REGION Network 333
   RUNG wire#powerrail
      Move(in := "DuplicateCarrierNumber", out1 => "Carrier_66_Duplicate_Carrier_Number")
   END_RUNG
   // the same network as SCL:
   "Carrier_66_Duplicate_Carrier_Number" := "DuplicateCarrierNumber";
END_REGION

REGION Network 334
   RUNG wire#powerrail
      Move(in := "FirstDuplicateCarrierPosition", out1 => "Carrier_66_First_Duplicate_Carrier_Position")
   END_RUNG
   // the same network as SCL:
   "Carrier_66_First_Duplicate_Carrier_Position" := "FirstDuplicateCarrierPosition";
END_REGION

REGION Network 335
   RUNG wire#powerrail
      Move(in := "SecondDuplicateCarrierPosition", out1 => "Carrier_66_Second_Duplicate_Carrier_Position")
   END_RUNG
   // the same network as SCL:
   "Carrier_66_Second_Duplicate_Carrier_Position" := "SecondDuplicateCarrierPosition";
END_REGION

REGION Network 336
   RUNG wire#powerrail
      Contact( "EMS".Carrier[66].SDC_OUT.HeartBeat )
      Coil( "Carrier_66_Heartbeat" )
   END_RUNG
   // the same network as SCL:
   "Carrier_66_Heartbeat" := "EMS".Carrier[66].SDC_OUT.HeartBeat;
END_REGION

REGION Network 337
   RUNG wire#powerrail
      Contact( "EMS".Carrier[66].SDC_OUT.DriveFwdCMD )
      I_Contact( "EMS".Carrier[65].SDC_IN.CrashDetectStatus )
      Coil( "Carrier_66_Drive_Forward_Command" )
   END_RUNG
   // the same network as SCL:
   "Carrier_66_Drive_Forward_Command" := "EMS".Carrier[66].SDC_OUT.DriveFwdCMD AND NOT "EMS".Carrier[65].SDC_IN.CrashDetectStatus;
END_REGION

REGION Network 338
   RUNG wire#powerrail
      Contact( "EMS".Carrier[66].SDC_OUT.FaultReset )
      Coil( "Carrier_66_Fault_Reset" )
   END_RUNG
   // the same network as SCL:
   "Carrier_66_Fault_Reset" := "EMS".Carrier[66].SDC_OUT.FaultReset;
END_REGION

REGION Network 339
   RUNG wire#powerrail
      Contact( "EMS".Carrier[66].SDC_OUT.AtCmdPos )
      Coil( "Carrier_66_At_Command_Position" )
   END_RUNG
   // the same network as SCL:
   "Carrier_66_At_Command_Position" := "EMS".Carrier[66].SDC_OUT.AtCmdPos;
END_REGION

REGION Network 340
   RUNG wire#powerrail
      Contact( "DuplicateCarrierfound" )
      Coil( "Carrier_66_Duplicate_Carrier_Fault" )
   END_RUNG
   // the same network as SCL:
   "Carrier_66_Duplicate_Carrier_Fault" := "DuplicateCarrierfound";
END_REGION

REGION Network 341
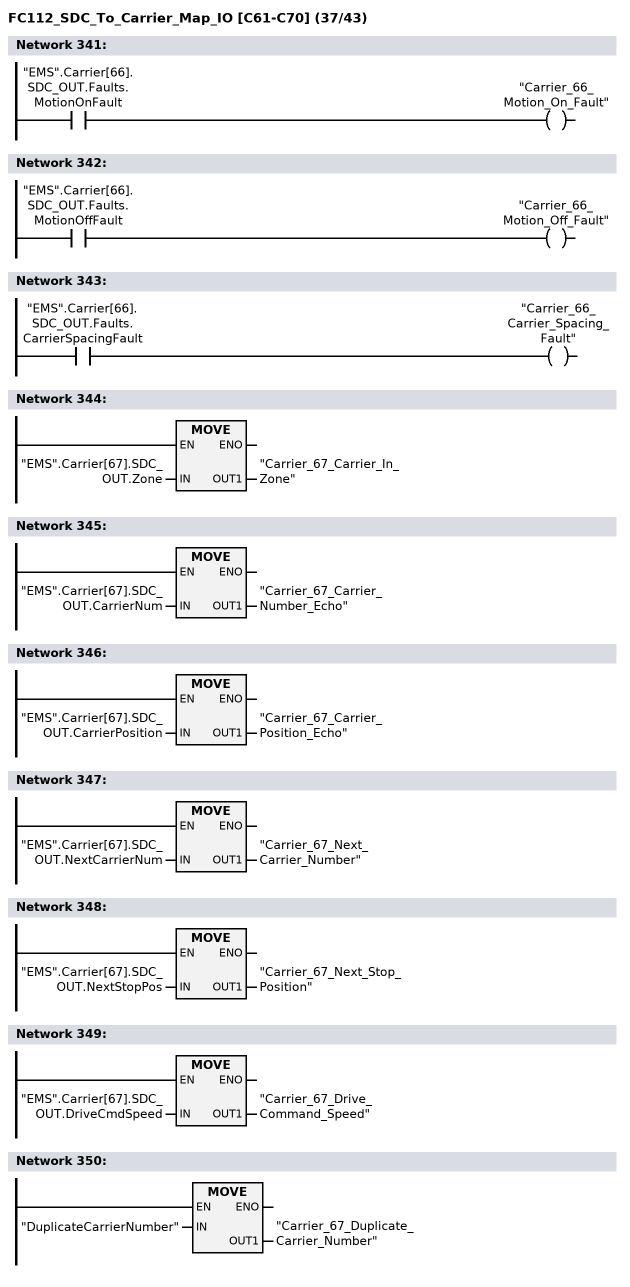
   RUNG wire#powerrail
      Contact( "EMS".Carrier[66].SDC_OUT.Faults.MotionOnFault )
      Coil( "Carrier_66_Motion_On_Fault" )
   END_RUNG
   // the same network as SCL:
   "Carrier_66_Motion_On_Fault" := "EMS".Carrier[66].SDC_OUT.Faults.MotionOnFault;
END_REGION

REGION Network 342
   RUNG wire#powerrail
      Contact( "EMS".Carrier[66].SDC_OUT.Faults.MotionOffFault )
      Coil( "Carrier_66_Motion_Off_Fault" )
   END_RUNG
   // the same network as SCL:
   "Carrier_66_Motion_Off_Fault" := "EMS".Carrier[66].SDC_OUT.Faults.MotionOffFault;
END_REGION

REGION Network 343
   RUNG wire#powerrail
      Contact( "EMS".Carrier[66].SDC_OUT.Faults.CarrierSpacingFault )
      Coil( "Carrier_66_Carrier_Spacing_Fault" )
   END_RUNG
   // the same network as SCL:
   "Carrier_66_Carrier_Spacing_Fault" := "EMS".Carrier[66].SDC_OUT.Faults.CarrierSpacingFault;
END_REGION

REGION Network 344
   RUNG wire#powerrail
      Move(in := "EMS".Carrier[67].SDC_OUT.Zone, out1 => "Carrier_67_Carrier_In_Zone")
   END_RUNG
   // the same network as SCL:
   "Carrier_67_Carrier_In_Zone" := "EMS".Carrier[67].SDC_OUT.Zone;
END_REGION

REGION Network 345
   RUNG wire#powerrail
      Move(in := "EMS".Carrier[67].SDC_OUT.CarrierNum, out1 => "Carrier_67_Carrier_Number_Echo")
   END_RUNG
   // the same network as SCL:
   "Carrier_67_Carrier_Number_Echo" := "EMS".Carrier[67].SDC_OUT.CarrierNum;
END_REGION

REGION Network 346
   RUNG wire#powerrail
      Move(in := "EMS".Carrier[67].SDC_OUT.CarrierPosition, out1 => "Carrier_67_Carrier_Position_Echo")
   END_RUNG
   // the same network as SCL:
   "Carrier_67_Carrier_Position_Echo" := "EMS".Carrier[67].SDC_OUT.CarrierPosition;
END_REGION

REGION Network 347
   RUNG wire#powerrail
      Move(in := "EMS".Carrier[67].SDC_OUT.NextCarrierNum, out1 => "Carrier_67_Next_Carrier_Number")
   END_RUNG
   // the same network as SCL:
   "Carrier_67_Next_Carrier_Number" := "EMS".Carrier[67].SDC_OUT.NextCarrierNum;
END_REGION

REGION Network 348
   RUNG wire#powerrail
      Move(in := "EMS".Carrier[67].SDC_OUT.NextStopPos, out1 => "Carrier_67_Next_Stop_Position")
   END_RUNG
   // the same network as SCL:
   "Carrier_67_Next_Stop_Position" := "EMS".Carrier[67].SDC_OUT.NextStopPos;
END_REGION

REGION Network 349
   RUNG wire#powerrail
      Move(in := "EMS".Carrier[67].SDC_OUT.DriveCmdSpeed, out1 => "Carrier_67_Drive_Command_Speed")
   END_RUNG
   // the same network as SCL:
   "Carrier_67_Drive_Command_Speed" := "EMS".Carrier[67].SDC_OUT.DriveCmdSpeed;
END_REGION

REGION Network 350
   RUNG wire#powerrail
      Move(in := "DuplicateCarrierNumber", out1 => "Carrier_67_Duplicate_Carrier_Number")
   END_RUNG
   // the same network as SCL:
   "Carrier_67_Duplicate_Carrier_Number" := "DuplicateCarrierNumber";
END_REGION

REGION Network 351
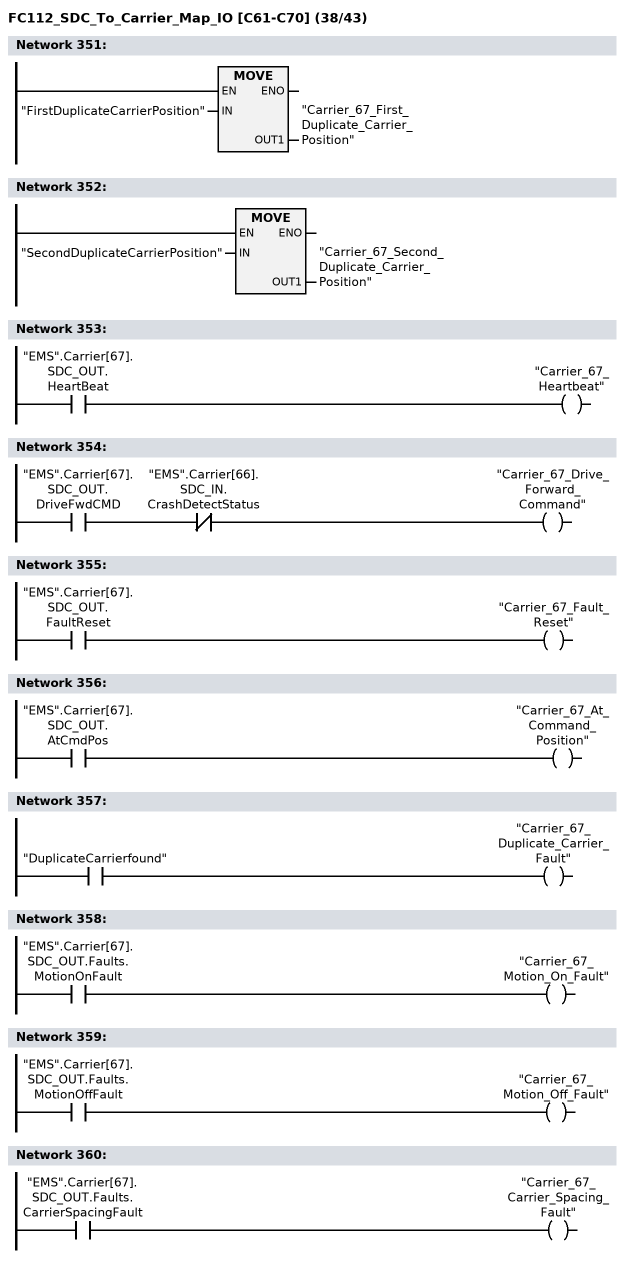
   RUNG wire#powerrail
      Move(in := "FirstDuplicateCarrierPosition", out1 => "Carrier_67_First_Duplicate_Carrier_Position")
   END_RUNG
   // the same network as SCL:
   "Carrier_67_First_Duplicate_Carrier_Position" := "FirstDuplicateCarrierPosition";
END_REGION

REGION Network 352
   RUNG wire#powerrail
      Move(in := "SecondDuplicateCarrierPosition", out1 => "Carrier_67_Second_Duplicate_Carrier_Position")
   END_RUNG
   // the same network as SCL:
   "Carrier_67_Second_Duplicate_Carrier_Position" := "SecondDuplicateCarrierPosition";
END_REGION

REGION Network 353
   RUNG wire#powerrail
      Contact( "EMS".Carrier[67].SDC_OUT.HeartBeat )
      Coil( "Carrier_67_Heartbeat" )
   END_RUNG
   // the same network as SCL:
   "Carrier_67_Heartbeat" := "EMS".Carrier[67].SDC_OUT.HeartBeat;
END_REGION

REGION Network 354
   RUNG wire#powerrail
      Contact( "EMS".Carrier[67].SDC_OUT.DriveFwdCMD )
      I_Contact( "EMS".Carrier[66].SDC_IN.CrashDetectStatus )
      Coil( "Carrier_67_Drive_Forward_Command" )
   END_RUNG
   // the same network as SCL:
   "Carrier_67_Drive_Forward_Command" := "EMS".Carrier[67].SDC_OUT.DriveFwdCMD AND NOT "EMS".Carrier[66].SDC_IN.CrashDetectStatus;
END_REGION

REGION Network 355
   RUNG wire#powerrail
      Contact( "EMS".Carrier[67].SDC_OUT.FaultReset )
      Coil( "Carrier_67_Fault_Reset" )
   END_RUNG
   // the same network as SCL:
   "Carrier_67_Fault_Reset" := "EMS".Carrier[67].SDC_OUT.FaultReset;
END_REGION

REGION Network 356
   RUNG wire#powerrail
      Contact( "EMS".Carrier[67].SDC_OUT.AtCmdPos )
      Coil( "Carrier_67_At_Command_Position" )
   END_RUNG
   // the same network as SCL:
   "Carrier_67_At_Command_Position" := "EMS".Carrier[67].SDC_OUT.AtCmdPos;
END_REGION

REGION Network 357
   RUNG wire#powerrail
      Contact( "DuplicateCarrierfound" )
      Coil( "Carrier_67_Duplicate_Carrier_Fault" )
   END_RUNG
   // the same network as SCL:
   "Carrier_67_Duplicate_Carrier_Fault" := "DuplicateCarrierfound";
END_REGION

REGION Network 358
   RUNG wire#powerrail
      Contact( "EMS".Carrier[67].SDC_OUT.Faults.MotionOnFault )
      Coil( "Carrier_67_Motion_On_Fault" )
   END_RUNG
   // the same network as SCL:
   "Carrier_67_Motion_On_Fault" := "EMS".Carrier[67].SDC_OUT.Faults.MotionOnFault;
END_REGION

REGION Network 359
   RUNG wire#powerrail
      Contact( "EMS".Carrier[67].SDC_OUT.Faults.MotionOffFault )
      Coil( "Carrier_67_Motion_Off_Fault" )
   END_RUNG
   // the same network as SCL:
   "Carrier_67_Motion_Off_Fault" := "EMS".Carrier[67].SDC_OUT.Faults.MotionOffFault;
END_REGION

REGION Network 360
   RUNG wire#powerrail
      Contact( "EMS".Carrier[67].SDC_OUT.Faults.CarrierSpacingFault )
      Coil( "Carrier_67_Carrier_Spacing_Fault" )
   END_RUNG
   // the same network as SCL:
   "Carrier_67_Carrier_Spacing_Fault" := "EMS".Carrier[67].SDC_OUT.Faults.CarrierSpacingFault;
END_REGION

REGION Network 361
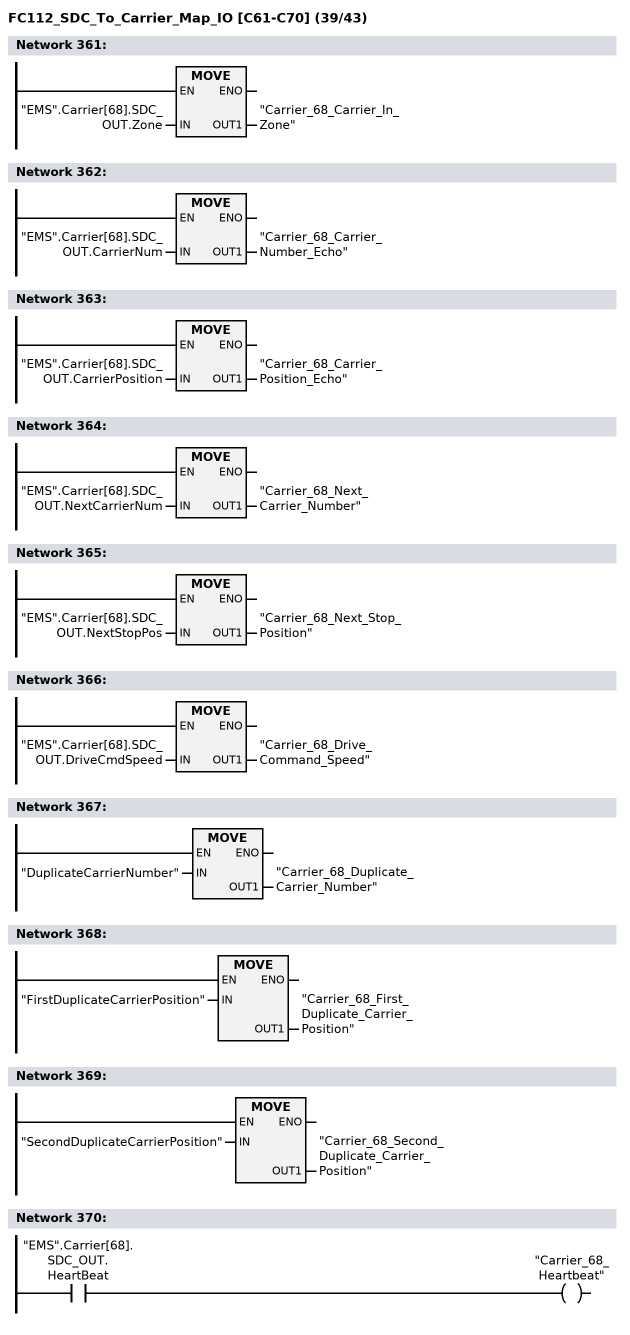
   RUNG wire#powerrail
      Move(in := "EMS".Carrier[68].SDC_OUT.Zone, out1 => "Carrier_68_Carrier_In_Zone")
   END_RUNG
   // the same network as SCL:
   "Carrier_68_Carrier_In_Zone" := "EMS".Carrier[68].SDC_OUT.Zone;
END_REGION

REGION Network 362
   RUNG wire#powerrail
      Move(in := "EMS".Carrier[68].SDC_OUT.CarrierNum, out1 => "Carrier_68_Carrier_Number_Echo")
   END_RUNG
   // the same network as SCL:
   "Carrier_68_Carrier_Number_Echo" := "EMS".Carrier[68].SDC_OUT.CarrierNum;
END_REGION

REGION Network 363
   RUNG wire#powerrail
      Move(in := "EMS".Carrier[68].SDC_OUT.CarrierPosition, out1 => "Carrier_68_Carrier_Position_Echo")
   END_RUNG
   // the same network as SCL:
   "Carrier_68_Carrier_Position_Echo" := "EMS".Carrier[68].SDC_OUT.CarrierPosition;
END_REGION

REGION Network 364
   RUNG wire#powerrail
      Move(in := "EMS".Carrier[68].SDC_OUT.NextCarrierNum, out1 => "Carrier_68_Next_Carrier_Number")
   END_RUNG
   // the same network as SCL:
   "Carrier_68_Next_Carrier_Number" := "EMS".Carrier[68].SDC_OUT.NextCarrierNum;
END_REGION

REGION Network 365
   RUNG wire#powerrail
      Move(in := "EMS".Carrier[68].SDC_OUT.NextStopPos, out1 => "Carrier_68_Next_Stop_Position")
   END_RUNG
   // the same network as SCL:
   "Carrier_68_Next_Stop_Position" := "EMS".Carrier[68].SDC_OUT.NextStopPos;
END_REGION

REGION Network 366
   RUNG wire#powerrail
      Move(in := "EMS".Carrier[68].SDC_OUT.DriveCmdSpeed, out1 => "Carrier_68_Drive_Command_Speed")
   END_RUNG
   // the same network as SCL:
   "Carrier_68_Drive_Command_Speed" := "EMS".Carrier[68].SDC_OUT.DriveCmdSpeed;
END_REGION

REGION Network 367
   RUNG wire#powerrail
      Move(in := "DuplicateCarrierNumber", out1 => "Carrier_68_Duplicate_Carrier_Number")
   END_RUNG
   // the same network as SCL:
   "Carrier_68_Duplicate_Carrier_Number" := "DuplicateCarrierNumber";
END_REGION

REGION Network 368
   RUNG wire#powerrail
      Move(in := "FirstDuplicateCarrierPosition", out1 => "Carrier_68_First_Duplicate_Carrier_Position")
   END_RUNG
   // the same network as SCL:
   "Carrier_68_First_Duplicate_Carrier_Position" := "FirstDuplicateCarrierPosition";
END_REGION

REGION Network 369
   RUNG wire#powerrail
      Move(in := "SecondDuplicateCarrierPosition", out1 => "Carrier_68_Second_Duplicate_Carrier_Position")
   END_RUNG
   // the same network as SCL:
   "Carrier_68_Second_Duplicate_Carrier_Position" := "SecondDuplicateCarrierPosition";
END_REGION

REGION Network 370
   RUNG wire#powerrail
      Contact( "EMS".Carrier[68].SDC_OUT.HeartBeat )
      Coil( "Carrier_68_Heartbeat" )
   END_RUNG
   // the same network as SCL:
   "Carrier_68_Heartbeat" := "EMS".Carrier[68].SDC_OUT.HeartBeat;
END_REGION

REGION Network 371
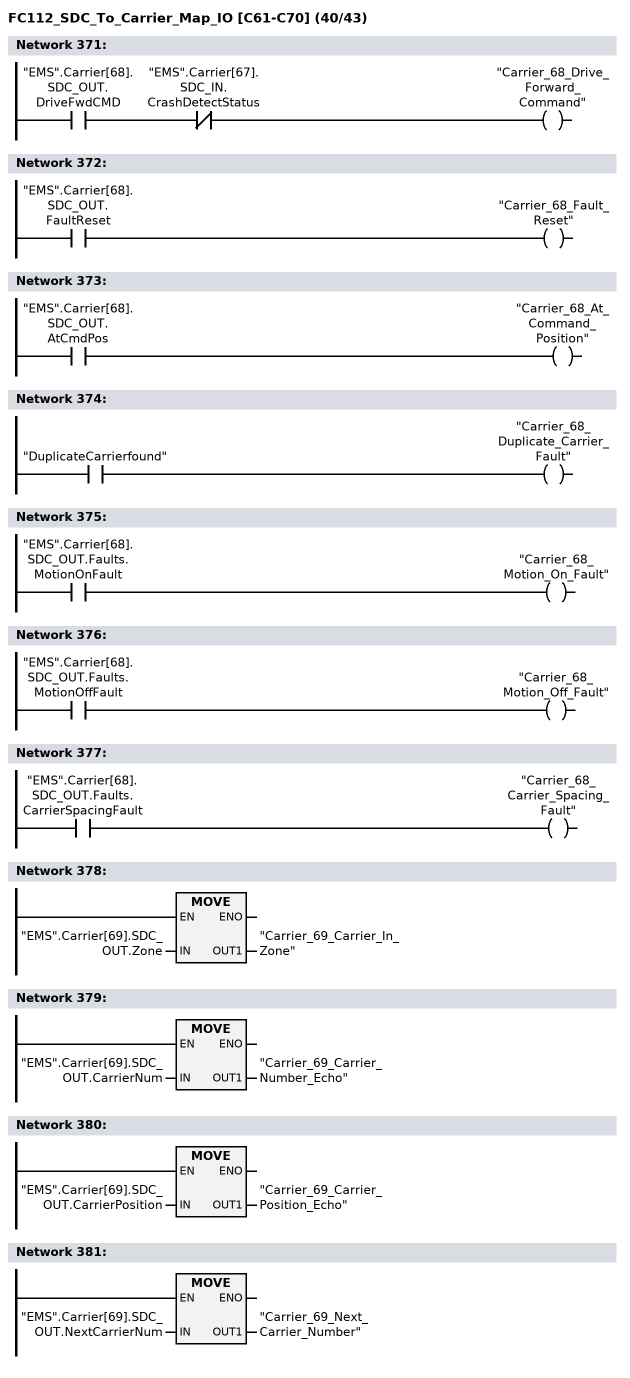
   RUNG wire#powerrail
      Contact( "EMS".Carrier[68].SDC_OUT.DriveFwdCMD )
      I_Contact( "EMS".Carrier[67].SDC_IN.CrashDetectStatus )
      Coil( "Carrier_68_Drive_Forward_Command" )
   END_RUNG
   // the same network as SCL:
   "Carrier_68_Drive_Forward_Command" := "EMS".Carrier[68].SDC_OUT.DriveFwdCMD AND NOT "EMS".Carrier[67].SDC_IN.CrashDetectStatus;
END_REGION

REGION Network 372
   RUNG wire#powerrail
      Contact( "EMS".Carrier[68].SDC_OUT.FaultReset )
      Coil( "Carrier_68_Fault_Reset" )
   END_RUNG
   // the same network as SCL:
   "Carrier_68_Fault_Reset" := "EMS".Carrier[68].SDC_OUT.FaultReset;
END_REGION

REGION Network 373
   RUNG wire#powerrail
      Contact( "EMS".Carrier[68].SDC_OUT.AtCmdPos )
      Coil( "Carrier_68_At_Command_Position" )
   END_RUNG
   // the same network as SCL:
   "Carrier_68_At_Command_Position" := "EMS".Carrier[68].SDC_OUT.AtCmdPos;
END_REGION

REGION Network 374
   RUNG wire#powerrail
      Contact( "DuplicateCarrierfound" )
      Coil( "Carrier_68_Duplicate_Carrier_Fault" )
   END_RUNG
   // the same network as SCL:
   "Carrier_68_Duplicate_Carrier_Fault" := "DuplicateCarrierfound";
END_REGION

REGION Network 375
   RUNG wire#powerrail
      Contact( "EMS".Carrier[68].SDC_OUT.Faults.MotionOnFault )
      Coil( "Carrier_68_Motion_On_Fault" )
   END_RUNG
   // the same network as SCL:
   "Carrier_68_Motion_On_Fault" := "EMS".Carrier[68].SDC_OUT.Faults.MotionOnFault;
END_REGION

REGION Network 376
   RUNG wire#powerrail
      Contact( "EMS".Carrier[68].SDC_OUT.Faults.MotionOffFault )
      Coil( "Carrier_68_Motion_Off_Fault" )
   END_RUNG
   // the same network as SCL:
   "Carrier_68_Motion_Off_Fault" := "EMS".Carrier[68].SDC_OUT.Faults.MotionOffFault;
END_REGION

REGION Network 377
   RUNG wire#powerrail
      Contact( "EMS".Carrier[68].SDC_OUT.Faults.CarrierSpacingFault )
      Coil( "Carrier_68_Carrier_Spacing_Fault" )
   END_RUNG
   // the same network as SCL:
   "Carrier_68_Carrier_Spacing_Fault" := "EMS".Carrier[68].SDC_OUT.Faults.CarrierSpacingFault;
END_REGION

REGION Network 378
   RUNG wire#powerrail
      Move(in := "EMS".Carrier[69].SDC_OUT.Zone, out1 => "Carrier_69_Carrier_In_Zone")
   END_RUNG
   // the same network as SCL:
   "Carrier_69_Carrier_In_Zone" := "EMS".Carrier[69].SDC_OUT.Zone;
END_REGION

REGION Network 379
   RUNG wire#powerrail
      Move(in := "EMS".Carrier[69].SDC_OUT.CarrierNum, out1 => "Carrier_69_Carrier_Number_Echo")
   END_RUNG
   // the same network as SCL:
   "Carrier_69_Carrier_Number_Echo" := "EMS".Carrier[69].SDC_OUT.CarrierNum;
END_REGION

REGION Network 380
   RUNG wire#powerrail
      Move(in := "EMS".Carrier[69].SDC_OUT.CarrierPosition, out1 => "Carrier_69_Carrier_Position_Echo")
   END_RUNG
   // the same network as SCL:
   "Carrier_69_Carrier_Position_Echo" := "EMS".Carrier[69].SDC_OUT.CarrierPosition;
END_REGION

REGION Network 381
   RUNG wire#powerrail
      Move(in := "EMS".Carrier[69].SDC_OUT.NextCarrierNum, out1 => "Carrier_69_Next_Carrier_Number")
   END_RUNG
   // the same network as SCL:
   "Carrier_69_Next_Carrier_Number" := "EMS".Carrier[69].SDC_OUT.NextCarrierNum;
END_REGION

REGION Network 382
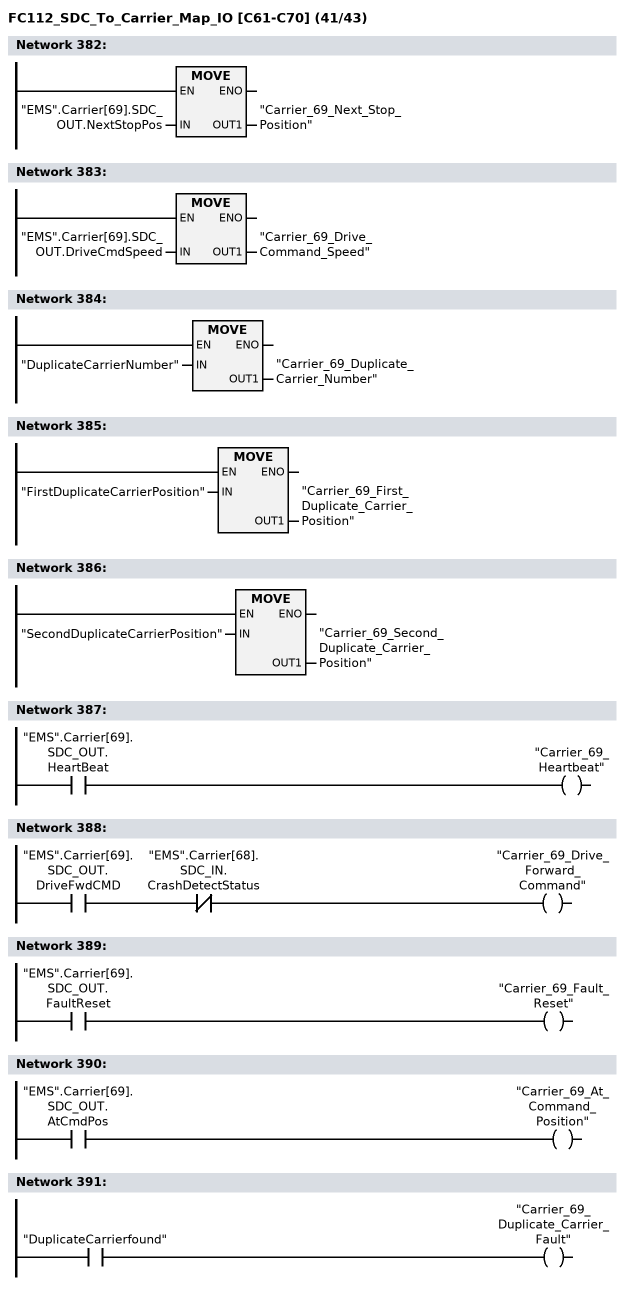
   RUNG wire#powerrail
      Move(in := "EMS".Carrier[69].SDC_OUT.NextStopPos, out1 => "Carrier_69_Next_Stop_Position")
   END_RUNG
   // the same network as SCL:
   "Carrier_69_Next_Stop_Position" := "EMS".Carrier[69].SDC_OUT.NextStopPos;
END_REGION

REGION Network 383
   RUNG wire#powerrail
      Move(in := "EMS".Carrier[69].SDC_OUT.DriveCmdSpeed, out1 => "Carrier_69_Drive_Command_Speed")
   END_RUNG
   // the same network as SCL:
   "Carrier_69_Drive_Command_Speed" := "EMS".Carrier[69].SDC_OUT.DriveCmdSpeed;
END_REGION

REGION Network 384
   RUNG wire#powerrail
      Move(in := "DuplicateCarrierNumber", out1 => "Carrier_69_Duplicate_Carrier_Number")
   END_RUNG
   // the same network as SCL:
   "Carrier_69_Duplicate_Carrier_Number" := "DuplicateCarrierNumber";
END_REGION

REGION Network 385
   RUNG wire#powerrail
      Move(in := "FirstDuplicateCarrierPosition", out1 => "Carrier_69_First_Duplicate_Carrier_Position")
   END_RUNG
   // the same network as SCL:
   "Carrier_69_First_Duplicate_Carrier_Position" := "FirstDuplicateCarrierPosition";
END_REGION

REGION Network 386
   RUNG wire#powerrail
      Move(in := "SecondDuplicateCarrierPosition", out1 => "Carrier_69_Second_Duplicate_Carrier_Position")
   END_RUNG
   // the same network as SCL:
   "Carrier_69_Second_Duplicate_Carrier_Position" := "SecondDuplicateCarrierPosition";
END_REGION

REGION Network 387
   RUNG wire#powerrail
      Contact( "EMS".Carrier[69].SDC_OUT.HeartBeat )
      Coil( "Carrier_69_Heartbeat" )
   END_RUNG
   // the same network as SCL:
   "Carrier_69_Heartbeat" := "EMS".Carrier[69].SDC_OUT.HeartBeat;
END_REGION

REGION Network 388
   RUNG wire#powerrail
      Contact( "EMS".Carrier[69].SDC_OUT.DriveFwdCMD )
      I_Contact( "EMS".Carrier[68].SDC_IN.CrashDetectStatus )
      Coil( "Carrier_69_Drive_Forward_Command" )
   END_RUNG
   // the same network as SCL:
   "Carrier_69_Drive_Forward_Command" := "EMS".Carrier[69].SDC_OUT.DriveFwdCMD AND NOT "EMS".Carrier[68].SDC_IN.CrashDetectStatus;
END_REGION

REGION Network 389
   RUNG wire#powerrail
      Contact( "EMS".Carrier[69].SDC_OUT.FaultReset )
      Coil( "Carrier_69_Fault_Reset" )
   END_RUNG
   // the same network as SCL:
   "Carrier_69_Fault_Reset" := "EMS".Carrier[69].SDC_OUT.FaultReset;
END_REGION

REGION Network 390
   RUNG wire#powerrail
      Contact( "EMS".Carrier[69].SDC_OUT.AtCmdPos )
      Coil( "Carrier_69_At_Command_Position" )
   END_RUNG
   // the same network as SCL:
   "Carrier_69_At_Command_Position" := "EMS".Carrier[69].SDC_OUT.AtCmdPos;
END_REGION

REGION Network 391
   RUNG wire#powerrail
      Contact( "DuplicateCarrierfound" )
      Coil( "Carrier_69_Duplicate_Carrier_Fault" )
   END_RUNG
   // the same network as SCL:
   "Carrier_69_Duplicate_Carrier_Fault" := "DuplicateCarrierfound";
END_REGION

REGION Network 392
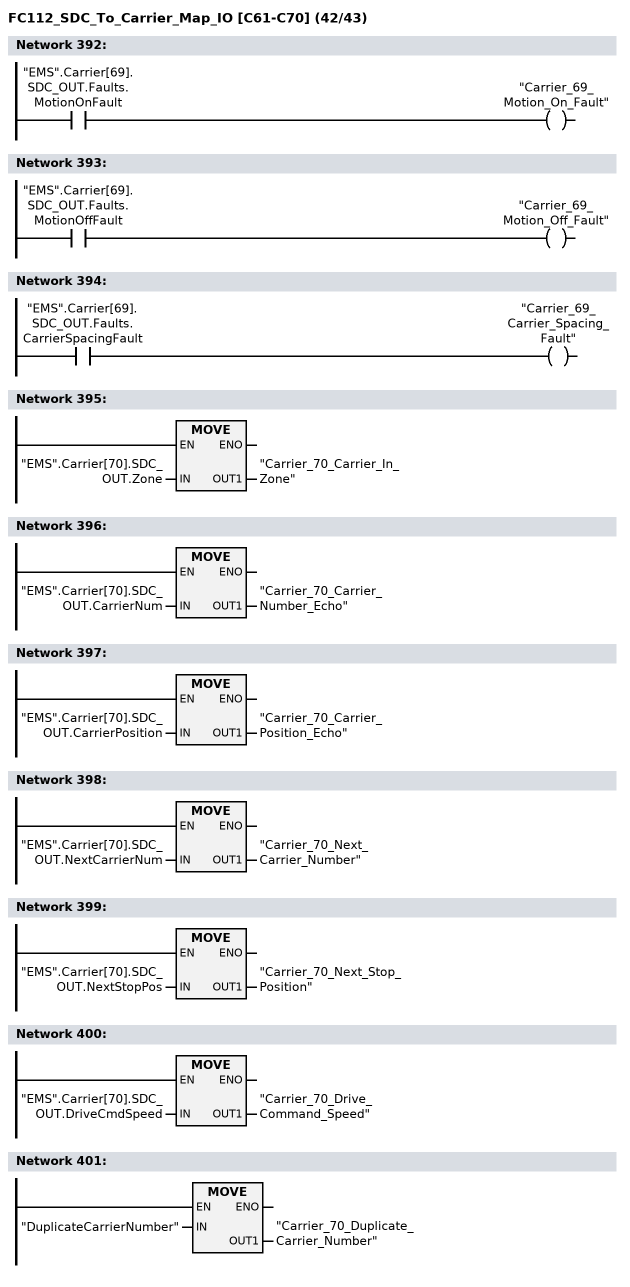
   RUNG wire#powerrail
      Contact( "EMS".Carrier[69].SDC_OUT.Faults.MotionOnFault )
      Coil( "Carrier_69_Motion_On_Fault" )
   END_RUNG
   // the same network as SCL:
   "Carrier_69_Motion_On_Fault" := "EMS".Carrier[69].SDC_OUT.Faults.MotionOnFault;
END_REGION

REGION Network 393
   RUNG wire#powerrail
      Contact( "EMS".Carrier[69].SDC_OUT.Faults.MotionOffFault )
      Coil( "Carrier_69_Motion_Off_Fault" )
   END_RUNG
   // the same network as SCL:
   "Carrier_69_Motion_Off_Fault" := "EMS".Carrier[69].SDC_OUT.Faults.MotionOffFault;
END_REGION

REGION Network 394
   RUNG wire#powerrail
      Contact( "EMS".Carrier[69].SDC_OUT.Faults.CarrierSpacingFault )
      Coil( "Carrier_69_Carrier_Spacing_Fault" )
   END_RUNG
   // the same network as SCL:
   "Carrier_69_Carrier_Spacing_Fault" := "EMS".Carrier[69].SDC_OUT.Faults.CarrierSpacingFault;
END_REGION

REGION Network 395
   RUNG wire#powerrail
      Move(in := "EMS".Carrier[70].SDC_OUT.Zone, out1 => "Carrier_70_Carrier_In_Zone")
   END_RUNG
   // the same network as SCL:
   "Carrier_70_Carrier_In_Zone" := "EMS".Carrier[70].SDC_OUT.Zone;
END_REGION

REGION Network 396
   RUNG wire#powerrail
      Move(in := "EMS".Carrier[70].SDC_OUT.CarrierNum, out1 => "Carrier_70_Carrier_Number_Echo")
   END_RUNG
   // the same network as SCL:
   "Carrier_70_Carrier_Number_Echo" := "EMS".Carrier[70].SDC_OUT.CarrierNum;
END_REGION

REGION Network 397
   RUNG wire#powerrail
      Move(in := "EMS".Carrier[70].SDC_OUT.CarrierPosition, out1 => "Carrier_70_Carrier_Position_Echo")
   END_RUNG
   // the same network as SCL:
   "Carrier_70_Carrier_Position_Echo" := "EMS".Carrier[70].SDC_OUT.CarrierPosition;
END_REGION

REGION Network 398
   RUNG wire#powerrail
      Move(in := "EMS".Carrier[70].SDC_OUT.NextCarrierNum, out1 => "Carrier_70_Next_Carrier_Number")
   END_RUNG
   // the same network as SCL:
   "Carrier_70_Next_Carrier_Number" := "EMS".Carrier[70].SDC_OUT.NextCarrierNum;
END_REGION

REGION Network 399
   RUNG wire#powerrail
      Move(in := "EMS".Carrier[70].SDC_OUT.NextStopPos, out1 => "Carrier_70_Next_Stop_Position")
   END_RUNG
   // the same network as SCL:
   "Carrier_70_Next_Stop_Position" := "EMS".Carrier[70].SDC_OUT.NextStopPos;
END_REGION

REGION Network 400
   RUNG wire#powerrail
      Move(in := "EMS".Carrier[70].SDC_OUT.DriveCmdSpeed, out1 => "Carrier_70_Drive_Command_Speed")
   END_RUNG
   // the same network as SCL:
   "Carrier_70_Drive_Command_Speed" := "EMS".Carrier[70].SDC_OUT.DriveCmdSpeed;
END_REGION

REGION Network 401
   RUNG wire#powerrail
      Move(in := "DuplicateCarrierNumber", out1 => "Carrier_70_Duplicate_Carrier_Number")
   END_RUNG
   // the same network as SCL:
   "Carrier_70_Duplicate_Carrier_Number" := "DuplicateCarrierNumber";
END_REGION

REGION Network 402
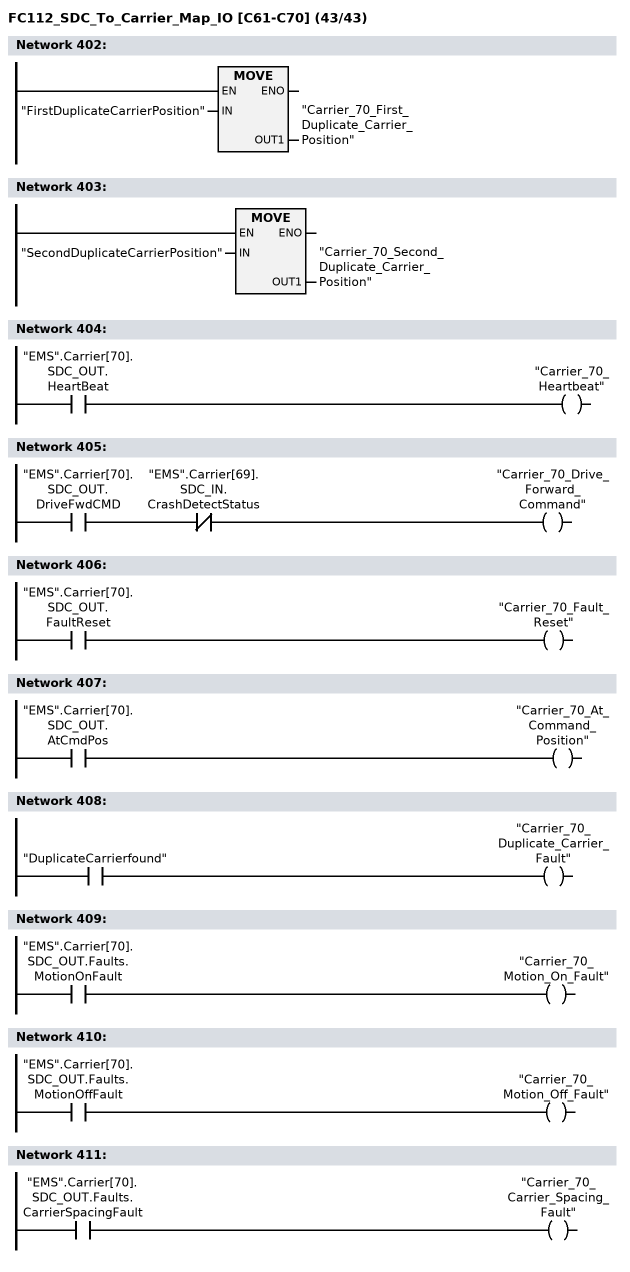
   RUNG wire#powerrail
      Move(in := "FirstDuplicateCarrierPosition", out1 => "Carrier_70_First_Duplicate_Carrier_Position")
   END_RUNG
   // the same network as SCL:
   "Carrier_70_First_Duplicate_Carrier_Position" := "FirstDuplicateCarrierPosition";
END_REGION

REGION Network 403
   RUNG wire#powerrail
      Move(in := "SecondDuplicateCarrierPosition", out1 => "Carrier_70_Second_Duplicate_Carrier_Position")
   END_RUNG
   // the same network as SCL:
   "Carrier_70_Second_Duplicate_Carrier_Position" := "SecondDuplicateCarrierPosition";
END_REGION

REGION Network 404
   RUNG wire#powerrail
      Contact( "EMS".Carrier[70].SDC_OUT.HeartBeat )
      Coil( "Carrier_70_Heartbeat" )
   END_RUNG
   // the same network as SCL:
   "Carrier_70_Heartbeat" := "EMS".Carrier[70].SDC_OUT.HeartBeat;
END_REGION

REGION Network 405
   RUNG wire#powerrail
      Contact( "EMS".Carrier[70].SDC_OUT.DriveFwdCMD )
      I_Contact( "EMS".Carrier[69].SDC_IN.CrashDetectStatus )
      Coil( "Carrier_70_Drive_Forward_Command" )
   END_RUNG
   // the same network as SCL:
   "Carrier_70_Drive_Forward_Command" := "EMS".Carrier[70].SDC_OUT.DriveFwdCMD AND NOT "EMS".Carrier[69].SDC_IN.CrashDetectStatus;
END_REGION

REGION Network 406
   RUNG wire#powerrail
      Contact( "EMS".Carrier[70].SDC_OUT.FaultReset )
      Coil( "Carrier_70_Fault_Reset" )
   END_RUNG
   // the same network as SCL:
   "Carrier_70_Fault_Reset" := "EMS".Carrier[70].SDC_OUT.FaultReset;
END_REGION

REGION Network 407
   RUNG wire#powerrail
      Contact( "EMS".Carrier[70].SDC_OUT.AtCmdPos )
      Coil( "Carrier_70_At_Command_Position" )
   END_RUNG
   // the same network as SCL:
   "Carrier_70_At_Command_Position" := "EMS".Carrier[70].SDC_OUT.AtCmdPos;
END_REGION

REGION Network 408
   RUNG wire#powerrail
      Contact( "DuplicateCarrierfound" )
      Coil( "Carrier_70_Duplicate_Carrier_Fault" )
   END_RUNG
   // the same network as SCL:
   "Carrier_70_Duplicate_Carrier_Fault" := "DuplicateCarrierfound";
END_REGION

REGION Network 409
   RUNG wire#powerrail
      Contact( "EMS".Carrier[70].SDC_OUT.Faults.MotionOnFault )
      Coil( "Carrier_70_Motion_On_Fault" )
   END_RUNG
   // the same network as SCL:
   "Carrier_70_Motion_On_Fault" := "EMS".Carrier[70].SDC_OUT.Faults.MotionOnFault;
END_REGION

REGION Network 410
   RUNG wire#powerrail
      Contact( "EMS".Carrier[70].SDC_OUT.Faults.MotionOffFault )
      Coil( "Carrier_70_Motion_Off_Fault" )
   END_RUNG
   // the same network as SCL:
   "Carrier_70_Motion_Off_Fault" := "EMS".Carrier[70].SDC_OUT.Faults.MotionOffFault;
END_REGION

REGION Network 411
   RUNG wire#powerrail
      Contact( "EMS".Carrier[70].SDC_OUT.Faults.CarrierSpacingFault )
      Coil( "Carrier_70_Carrier_Spacing_Fault" )
   END_RUNG
   // the same network as SCL:
   "Carrier_70_Carrier_Spacing_Fault" := "EMS".Carrier[70].SDC_OUT.Faults.CarrierSpacingFault;
END_REGION
END_FUNCTION

FUNCTION "FC113_SDC_To_Carrier_Map_IO [C71-C80]" : Void   // FC113, LAD
{ S7_Optimized_Access := 'TRUE' }
VERSION : 0.1
BEGIN

REGION Network 1
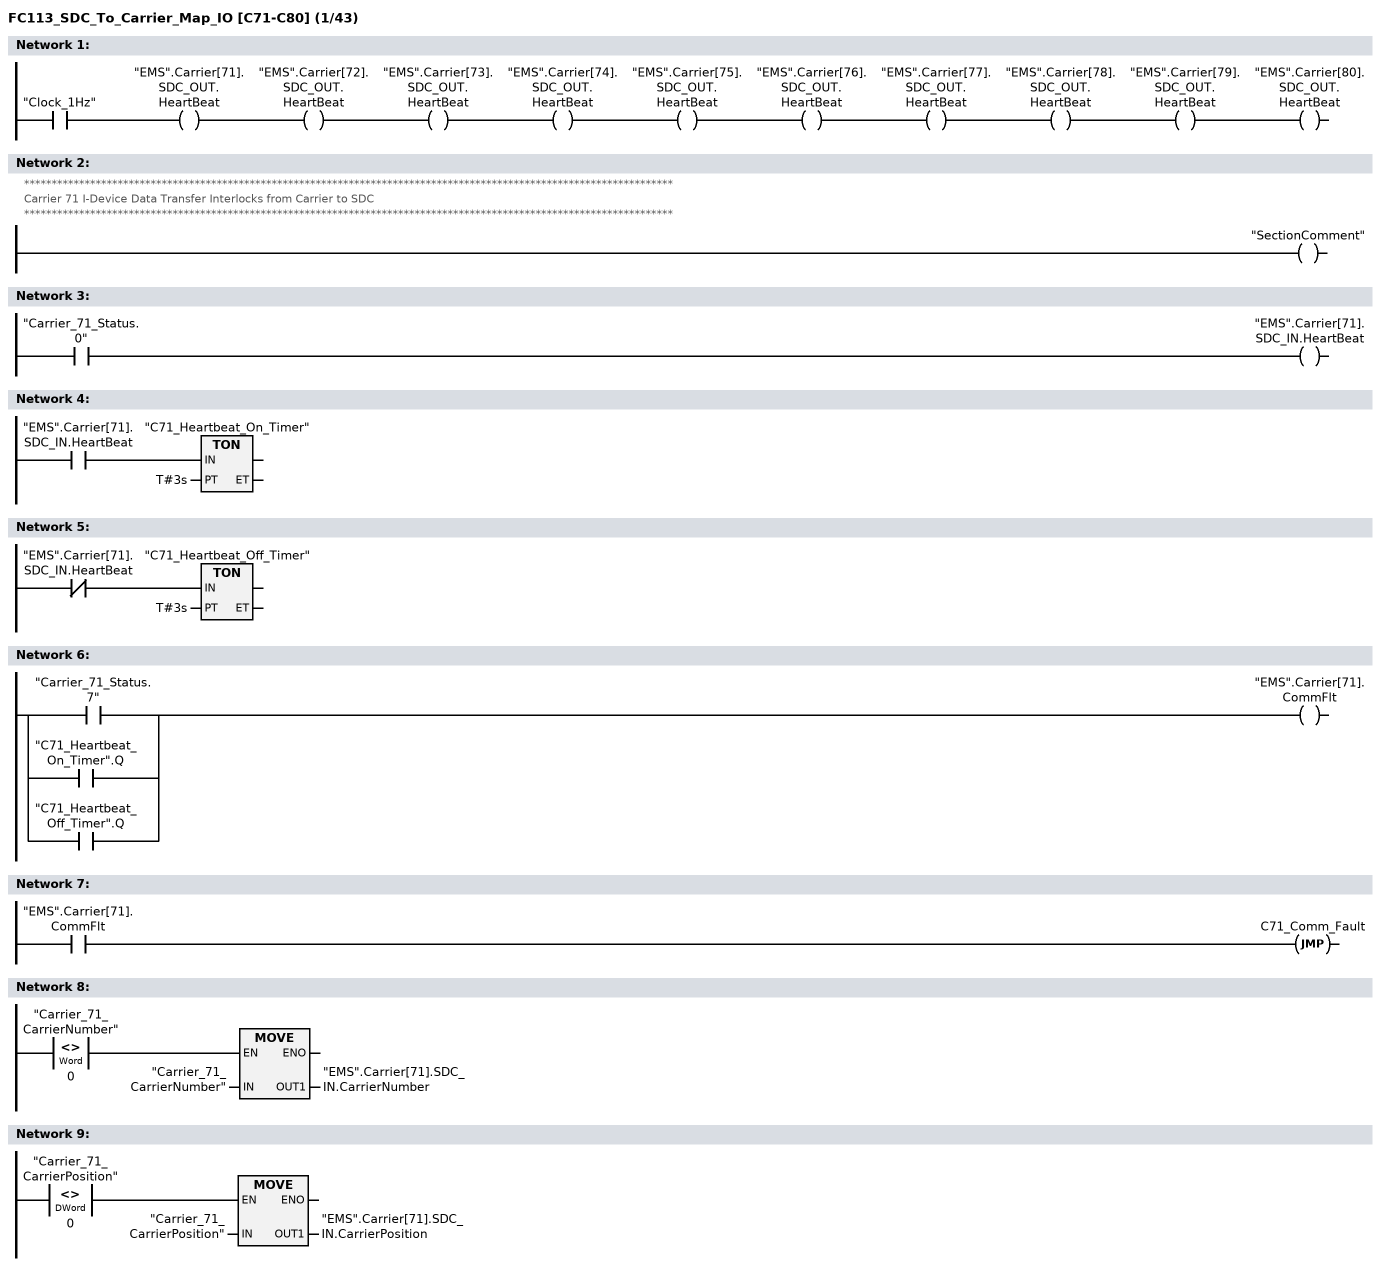
   RUNG wire#powerrail
      Contact( "Clock_1Hz" )
      Coil( "EMS".Carrier[71].SDC_OUT.HeartBeat )
      Coil( "EMS".Carrier[72].SDC_OUT.HeartBeat )
      Coil( "EMS".Carrier[73].SDC_OUT.HeartBeat )
      Coil( "EMS".Carrier[74].SDC_OUT.HeartBeat )
      Coil( "EMS".Carrier[75].SDC_OUT.HeartBeat )
      Coil( "EMS".Carrier[76].SDC_OUT.HeartBeat )
      Coil( "EMS".Carrier[77].SDC_OUT.HeartBeat )
      Coil( "EMS".Carrier[78].SDC_OUT.HeartBeat )
      Coil( "EMS".Carrier[79].SDC_OUT.HeartBeat )
      Coil( "EMS".Carrier[80].SDC_OUT.HeartBeat )
   END_RUNG
   // the same network as SCL:
   "EMS".Carrier[71].SDC_OUT.HeartBeat := "Clock_1Hz";
   "EMS".Carrier[72].SDC_OUT.HeartBeat := "Clock_1Hz";
   "EMS".Carrier[73].SDC_OUT.HeartBeat := "Clock_1Hz";
   "EMS".Carrier[74].SDC_OUT.HeartBeat := "Clock_1Hz";
   "EMS".Carrier[75].SDC_OUT.HeartBeat := "Clock_1Hz";
   "EMS".Carrier[76].SDC_OUT.HeartBeat := "Clock_1Hz";
   "EMS".Carrier[77].SDC_OUT.HeartBeat := "Clock_1Hz";